REGION Network 13: ENCENDIDO ACTUADORES TUNEL 1
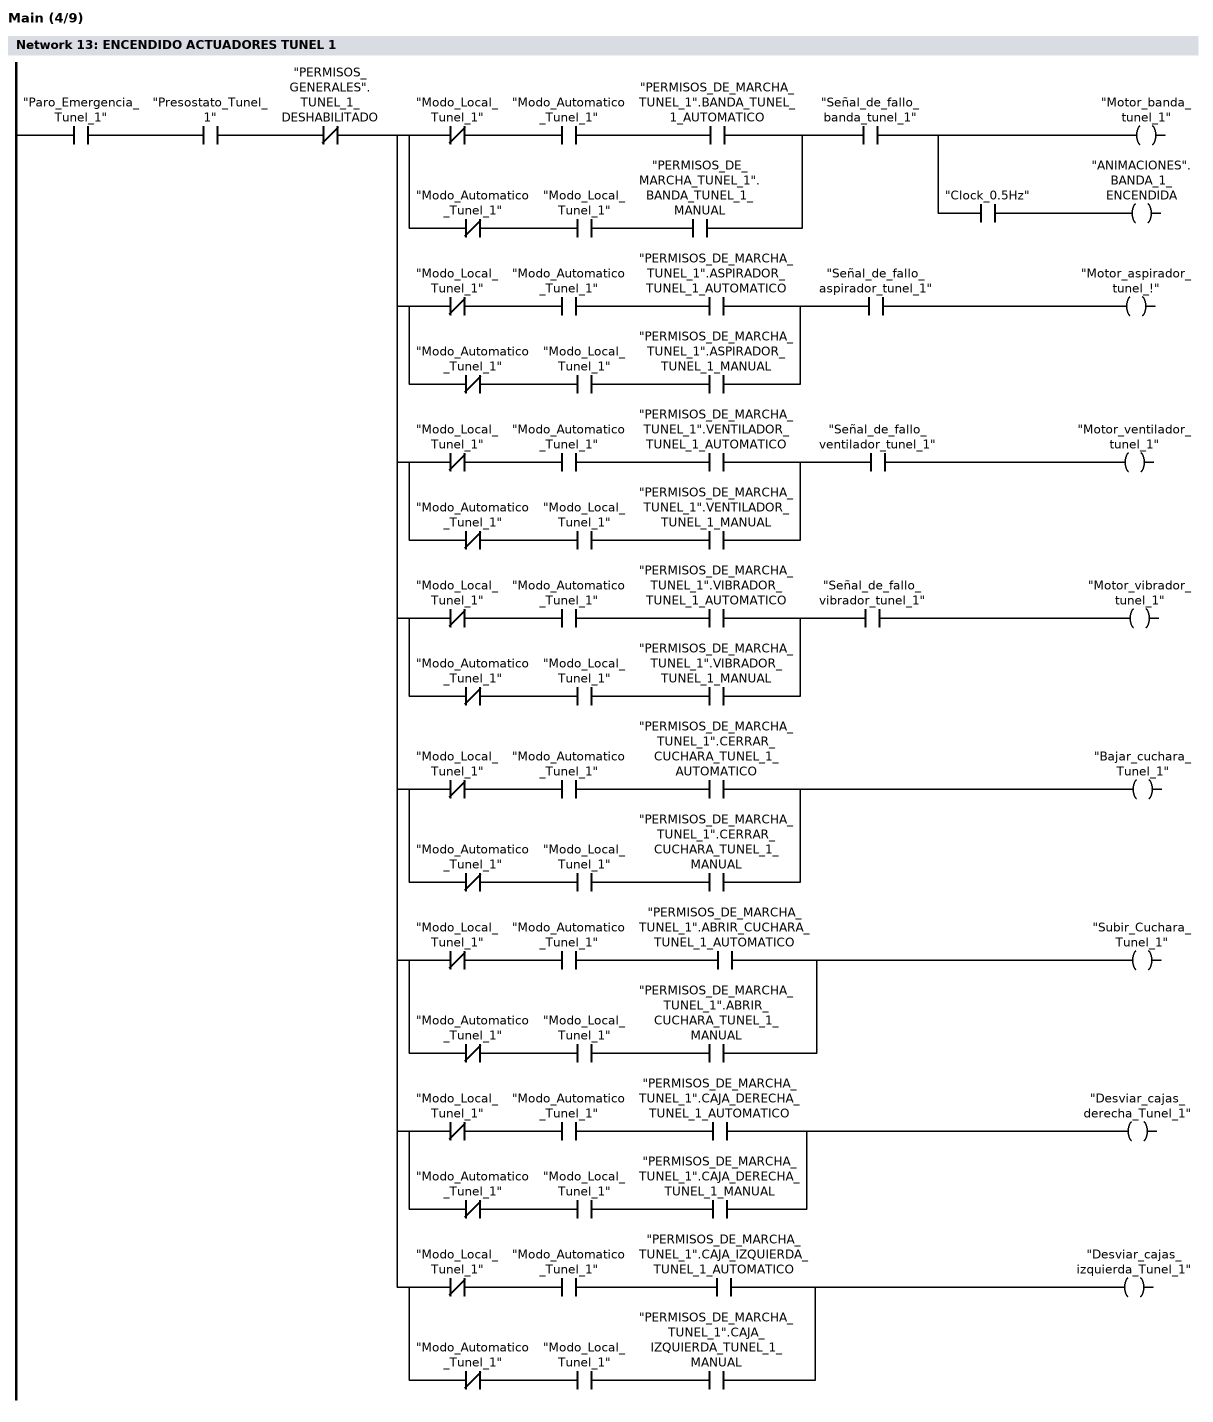
   RUNG wire#powerrail
      Contact( "Paro_Emergencia_Tunel_1" )
      Contact( "Presostato_Tunel_1" )
      I_Contact( "PERMISOS_GENERALES".TUNEL_1_DESHABILITADO )
      wire#w1
      I_Contact( "Modo_Local_Tunel_1" )
      Contact( "Modo_Automatico_Tunel_1" )
      Contact( "PERMISOS_DE_MARCHA_TUNEL_1".BANDA_TUNEL_1_AUTOMATICO )
      wire#w2
      Contact( "Señal_de_fallo_banda_tunel_1" )
      wire#w3
      Coil( "Motor_banda_tunel_1" )
   END_RUNG
   RUNG wire#w1
      I_Contact( "Modo_Automatico_Tunel_1" )
      Contact( "Modo_Local_Tunel_1" )
      Contact( "PERMISOS_DE_MARCHA_TUNEL_1".BANDA_TUNEL_1_MANUAL )
   END_RUNG wire#w2
   RUNG wire#w3
      Contact( "Clock_0.5Hz" )
      Coil( "ANIMACIONES".BANDA_1_ENCENDIDA )
   END_RUNG
   RUNG wire#w1
      I_Contact( "Modo_Local_Tunel_1" )
      Contact( "Modo_Automatico_Tunel_1" )
      Contact( "PERMISOS_DE_MARCHA_TUNEL_1".ASPIRADOR_TUNEL_1_AUTOMATICO )
      wire#w4
      Contact( "Señal_de_fallo_aspirador_tunel_1" )
      Coil( "Motor_aspirador_tunel_!" )
   END_RUNG
   RUNG wire#w1
      I_Contact( "Modo_Automatico_Tunel_1" )
      Contact( "Modo_Local_Tunel_1" )
      Contact( "PERMISOS_DE_MARCHA_TUNEL_1".ASPIRADOR_TUNEL_1_MANUAL )
   END_RUNG wire#w4
   RUNG wire#w1
      I_Contact( "Modo_Local_Tunel_1" )
      Contact( "Modo_Automatico_Tunel_1" )
      Contact( "PERMISOS_DE_MARCHA_TUNEL_1".VENTILADOR_TUNEL_1_AUTOMATICO )
      wire#w5
      Contact( "Señal_de_fallo_ventilador_tunel_1" )
      Coil( "Motor_ventilador_tunel_1" )
   END_RUNG
   RUNG wire#w1
      I_Contact( "Modo_Automatico_Tunel_1" )
      Contact( "Modo_Local_Tunel_1" )
      Contact( "PERMISOS_DE_MARCHA_TUNEL_1".VENTILADOR_TUNEL_1_MANUAL )
   END_RUNG wire#w5
   RUNG wire#w1
      I_Contact( "Modo_Local_Tunel_1" )
      Contact( "Modo_Automatico_Tunel_1" )
      Contact( "PERMISOS_DE_MARCHA_TUNEL_1".VIBRADOR_TUNEL_1_AUTOMATICO )
      wire#w6
      Contact( "Señal_de_fallo_vibrador_tunel_1" )
      Coil( "Motor_vibrador_tunel_1" )
   END_RUNG
   RUNG wire#w1
      I_Contact( "Modo_Automatico_Tunel_1" )
      Contact( "Modo_Local_Tunel_1" )
      Contact( "PERMISOS_DE_MARCHA_TUNEL_1".VIBRADOR_TUNEL_1_MANUAL )
   END_RUNG wire#w6
   RUNG wire#w1
      I_Contact( "Modo_Local_Tunel_1" )
      Contact( "Modo_Automatico_Tunel_1" )
      Contact( "PERMISOS_DE_MARCHA_TUNEL_1".CERRAR_CUCHARA_TUNEL_1_AUTOMATICO )
      wire#w7
      Coil( "Bajar_cuchara_Tunel_1" )
   END_RUNG
   RUNG wire#w1
      I_Contact( "Modo_Automatico_Tunel_1" )
      Contact( "Modo_Local_Tunel_1" )
      Contact( "PERMISOS_DE_MARCHA_TUNEL_1".CERRAR_CUCHARA_TUNEL_1_MANUAL )
   END_RUNG wire#w7
   RUNG wire#w1
      I_Contact( "Modo_Local_Tunel_1" )
      Contact( "Modo_Automatico_Tunel_1" )
      Contact( "PERMISOS_DE_MARCHA_TUNEL_1".ABRIR_CUCHARA_TUNEL_1_AUTOMATICO )
      wire#w8
      Coil( "Subir_Cuchara_Tunel_1" )
   END_RUNG
   RUNG wire#w1
      I_Contact( "Modo_Automatico_Tunel_1" )
      Contact( "Modo_Local_Tunel_1" )
      Contact( "PERMISOS_DE_MARCHA_TUNEL_1".ABRIR_CUCHARA_TUNEL_1_MANUAL )
   END_RUNG wire#w8
   RUNG wire#w1
      I_Contact( "Modo_Local_Tunel_1" )
      Contact( "Modo_Automatico_Tunel_1" )
      Contact( "PERMISOS_DE_MARCHA_TUNEL_1".CAJA_DERECHA_TUNEL_1_AUTOMATICO )
      wire#w9
      Coil( "Desviar_cajas_derecha_Tunel_1" )
   END_RUNG
   RUNG wire#w1
      I_Contact( "Modo_Automatico_Tunel_1" )
      Contact( "Modo_Local_Tunel_1" )
      Contact( "PERMISOS_DE_MARCHA_TUNEL_1".CAJA_DERECHA_TUNEL_1_MANUAL )
   END_RUNG wire#w9
   RUNG wire#w1
      I_Contact( "Modo_Local_Tunel_1" )
      Contact( "Modo_Automatico_Tunel_1" )
      Contact( "PERMISOS_DE_MARCHA_TUNEL_1".CAJA_IZQUIERDA_TUNEL_1_AUTOMATICO )
      wire#w10
      Coil( "Desviar_cajas_izquierda_Tunel_1" )
   END_RUNG
   RUNG wire#w1
      I_Contact( "Modo_Automatico_Tunel_1" )
      Contact( "Modo_Local_Tunel_1" )
      Contact( "PERMISOS_DE_MARCHA_TUNEL_1".CAJA_IZQUIERDA_TUNEL_1_MANUAL )
   END_RUNG wire#w10
   // the same network as SCL:
   #_w1 := "Paro_Emergencia_Tunel_1" AND "Presostato_Tunel_1" AND NOT "PERMISOS_GENERALES".TUNEL_1_DESHABILITADO;
   "Motor_banda_tunel_1" := #_w1 AND ((NOT "Modo_Local_Tunel_1" AND "Modo_Automatico_Tunel_1" AND "PERMISOS_DE_MARCHA_TUNEL_1".BANDA_TUNEL_1_AUTOMATICO) OR (NOT "Modo_Automatico_Tunel_1" AND "Modo_Local_Tunel_1" AND "PERMISOS_DE_MARCHA_TUNEL_1".BANDA_TUNEL_1_MANUAL)) AND "Señal_de_fallo_banda_tunel_1";
   "ANIMACIONES".BANDA_1_ENCENDIDA := "Motor_banda_tunel_1" AND "Clock_0.5Hz";
   "Motor_aspirador_tunel_!" := #_w1 AND ((NOT "Modo_Local_Tunel_1" AND "Modo_Automatico_Tunel_1" AND "PERMISOS_DE_MARCHA_TUNEL_1".ASPIRADOR_TUNEL_1_AUTOMATICO) OR (NOT "Modo_Automatico_Tunel_1" AND "Modo_Local_Tunel_1" AND "PERMISOS_DE_MARCHA_TUNEL_1".ASPIRADOR_TUNEL_1_MANUAL)) AND "Señal_de_fallo_aspirador_tunel_1";
   "Motor_ventilador_tunel_1" := #_w1 AND ((NOT "Modo_Local_Tunel_1" AND "Modo_Automatico_Tunel_1" AND "PERMISOS_DE_MARCHA_TUNEL_1".VENTILADOR_TUNEL_1_AUTOMATICO) OR (NOT "Modo_Automatico_Tunel_1" AND "Modo_Local_Tunel_1" AND "PERMISOS_DE_MARCHA_TUNEL_1".VENTILADOR_TUNEL_1_MANUAL)) AND "Señal_de_fallo_ventilador_tunel_1";
   "Motor_vibrador_tunel_1" := #_w1 AND ((NOT "Modo_Local_Tunel_1" AND "Modo_Automatico_Tunel_1" AND "PERMISOS_DE_MARCHA_TUNEL_1".VIBRADOR_TUNEL_1_AUTOMATICO) OR (NOT "Modo_Automatico_Tunel_1" AND "Modo_Local_Tunel_1" AND "PERMISOS_DE_MARCHA_TUNEL_1".VIBRADOR_TUNEL_1_MANUAL)) AND "Señal_de_fallo_vibrador_tunel_1";
   "Bajar_cuchara_Tunel_1" := #_w1 AND ((NOT "Modo_Local_Tunel_1" AND "Modo_Automatico_Tunel_1" AND "PERMISOS_DE_MARCHA_TUNEL_1".CERRAR_CUCHARA_TUNEL_1_AUTOMATICO) OR (NOT "Modo_Automatico_Tunel_1" AND "Modo_Local_Tunel_1" AND "PERMISOS_DE_MARCHA_TUNEL_1".CERRAR_CUCHARA_TUNEL_1_MANUAL));
   "Subir_Cuchara_Tunel_1" := #_w1 AND ((NOT "Modo_Local_Tunel_1" AND "Modo_Automatico_Tunel_1" AND "PERMISOS_DE_MARCHA_TUNEL_1".ABRIR_CUCHARA_TUNEL_1_AUTOMATICO) OR (NOT "Modo_Automatico_Tunel_1" AND "Modo_Local_Tunel_1" AND "PERMISOS_DE_MARCHA_TUNEL_1".ABRIR_CUCHARA_TUNEL_1_MANUAL));
   "Desviar_cajas_derecha_Tunel_1" := #_w1 AND ((NOT "Modo_Local_Tunel_1" AND "Modo_Automatico_Tunel_1" AND "PERMISOS_DE_MARCHA_TUNEL_1".CAJA_DERECHA_TUNEL_1_AUTOMATICO) OR (NOT "Modo_Automatico_Tunel_1" AND "Modo_Local_Tunel_1" AND "PERMISOS_DE_MARCHA_TUNEL_1".CAJA_DERECHA_TUNEL_1_MANUAL));
   "Desviar_cajas_izquierda_Tunel_1" := #_w1 AND ((NOT "Modo_Local_Tunel_1" AND "Modo_Automatico_Tunel_1" AND "PERMISOS_DE_MARCHA_TUNEL_1".CAJA_IZQUIERDA_TUNEL_1_AUTOMATICO) OR (NOT "Modo_Automatico_Tunel_1" AND "Modo_Local_Tunel_1" AND "PERMISOS_DE_MARCHA_TUNEL_1".CAJA_IZQUIERDA_TUNEL_1_MANUAL));
END_REGION

REGION Network 14: ENCENDIDO ACTUADORES TUNEL 2
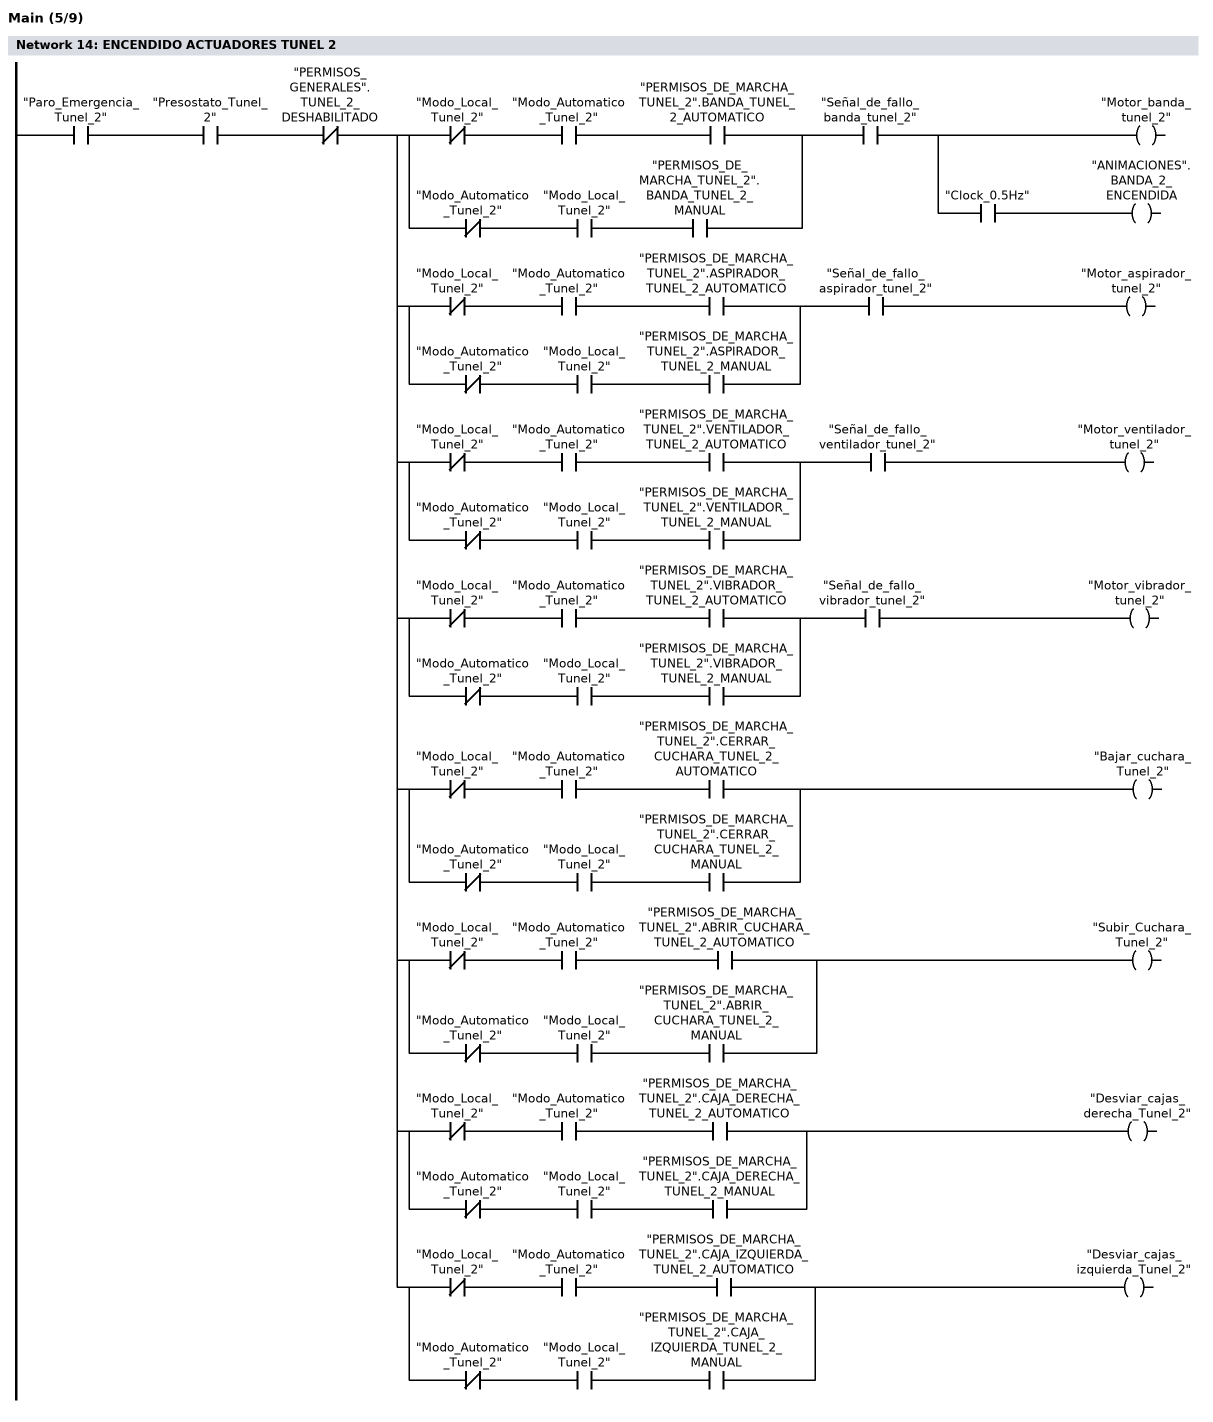
   RUNG wire#powerrail
      Contact( "Paro_Emergencia_Tunel_2" )
      Contact( "Presostato_Tunel_2" )
      I_Contact( "PERMISOS_GENERALES".TUNEL_2_DESHABILITADO )
      wire#w1
      I_Contact( "Modo_Local_Tunel_2" )
      Contact( "Modo_Automatico_Tunel_2" )
      Contact( "PERMISOS_DE_MARCHA_TUNEL_2".BANDA_TUNEL_2_AUTOMATICO )
      wire#w2
      Contact( "Señal_de_fallo_banda_tunel_2" )
      wire#w3
      Coil( "Motor_banda_tunel_2" )
   END_RUNG
   RUNG wire#w1
      I_Contact( "Modo_Automatico_Tunel_2" )
      Contact( "Modo_Local_Tunel_2" )
      Contact( "PERMISOS_DE_MARCHA_TUNEL_2".BANDA_TUNEL_2_MANUAL )
   END_RUNG wire#w2
   RUNG wire#w3
      Contact( "Clock_0.5Hz" )
      Coil( "ANIMACIONES".BANDA_2_ENCENDIDA )
   END_RUNG
   RUNG wire#w1
      I_Contact( "Modo_Local_Tunel_2" )
      Contact( "Modo_Automatico_Tunel_2" )
      Contact( "PERMISOS_DE_MARCHA_TUNEL_2".ASPIRADOR_TUNEL_2_AUTOMATICO )
      wire#w4
      Contact( "Señal_de_fallo_aspirador_tunel_2" )
      Coil( "Motor_aspirador_tunel_2" )
   END_RUNG
   RUNG wire#w1
      I_Contact( "Modo_Automatico_Tunel_2" )
      Contact( "Modo_Local_Tunel_2" )
      Contact( "PERMISOS_DE_MARCHA_TUNEL_2".ASPIRADOR_TUNEL_2_MANUAL )
   END_RUNG wire#w4
   RUNG wire#w1
      I_Contact( "Modo_Local_Tunel_2" )
      Contact( "Modo_Automatico_Tunel_2" )
      Contact( "PERMISOS_DE_MARCHA_TUNEL_2".VENTILADOR_TUNEL_2_AUTOMATICO )
      wire#w5
      Contact( "Señal_de_fallo_ventilador_tunel_2" )
      Coil( "Motor_ventilador_tunel_2" )
   END_RUNG
   RUNG wire#w1
      I_Contact( "Modo_Automatico_Tunel_2" )
      Contact( "Modo_Local_Tunel_2" )
      Contact( "PERMISOS_DE_MARCHA_TUNEL_2".VENTILADOR_TUNEL_2_MANUAL )
   END_RUNG wire#w5
   RUNG wire#w1
      I_Contact( "Modo_Local_Tunel_2" )
      Contact( "Modo_Automatico_Tunel_2" )
      Contact( "PERMISOS_DE_MARCHA_TUNEL_2".VIBRADOR_TUNEL_2_AUTOMATICO )
      wire#w6
      Contact( "Señal_de_fallo_vibrador_tunel_2" )
      Coil( "Motor_vibrador_tunel_2" )
   END_RUNG
   RUNG wire#w1
      I_Contact( "Modo_Automatico_Tunel_2" )
      Contact( "Modo_Local_Tunel_2" )
      Contact( "PERMISOS_DE_MARCHA_TUNEL_2".VIBRADOR_TUNEL_2_MANUAL )
   END_RUNG wire#w6
   RUNG wire#w1
      I_Contact( "Modo_Local_Tunel_2" )
      Contact( "Modo_Automatico_Tunel_2" )
      Contact( "PERMISOS_DE_MARCHA_TUNEL_2".CERRAR_CUCHARA_TUNEL_2_AUTOMATICO )
      wire#w7
      Coil( "Bajar_cuchara_Tunel_2" )
   END_RUNG
   RUNG wire#w1
      I_Contact( "Modo_Automatico_Tunel_2" )
      Contact( "Modo_Local_Tunel_2" )
      Contact( "PERMISOS_DE_MARCHA_TUNEL_2".CERRAR_CUCHARA_TUNEL_2_MANUAL )
   END_RUNG wire#w7
   RUNG wire#w1
      I_Contact( "Modo_Local_Tunel_2" )
      Contact( "Modo_Automatico_Tunel_2" )
      Contact( "PERMISOS_DE_MARCHA_TUNEL_2".ABRIR_CUCHARA_TUNEL_2_AUTOMATICO )
      wire#w8
      Coil( "Subir_Cuchara_Tunel_2" )
   END_RUNG
   RUNG wire#w1
      I_Contact( "Modo_Automatico_Tunel_2" )
      Contact( "Modo_Local_Tunel_2" )
      Contact( "PERMISOS_DE_MARCHA_TUNEL_2".ABRIR_CUCHARA_TUNEL_2_MANUAL )
   END_RUNG wire#w8
   RUNG wire#w1
      I_Contact( "Modo_Local_Tunel_2" )
      Contact( "Modo_Automatico_Tunel_2" )
      Contact( "PERMISOS_DE_MARCHA_TUNEL_2".CAJA_DERECHA_TUNEL_2_AUTOMATICO )
      wire#w9
      Coil( "Desviar_cajas_derecha_Tunel_2" )
   END_RUNG
   RUNG wire#w1
      I_Contact( "Modo_Automatico_Tunel_2" )
      Contact( "Modo_Local_Tunel_2" )
      Contact( "PERMISOS_DE_MARCHA_TUNEL_2".CAJA_DERECHA_TUNEL_2_MANUAL )
   END_RUNG wire#w9
   RUNG wire#w1
      I_Contact( "Modo_Local_Tunel_2" )
      Contact( "Modo_Automatico_Tunel_2" )
      Contact( "PERMISOS_DE_MARCHA_TUNEL_2".CAJA_IZQUIERDA_TUNEL_2_AUTOMATICO )
      wire#w10
      Coil( "Desviar_cajas_izquierda_Tunel_2" )
   END_RUNG
   RUNG wire#w1
      I_Contact( "Modo_Automatico_Tunel_2" )
      Contact( "Modo_Local_Tunel_2" )
      Contact( "PERMISOS_DE_MARCHA_TUNEL_2".CAJA_IZQUIERDA_TUNEL_2_MANUAL )
   END_RUNG wire#w10
   // the same network as SCL:
   #_w1 := "Paro_Emergencia_Tunel_2" AND "Presostato_Tunel_2" AND NOT "PERMISOS_GENERALES".TUNEL_2_DESHABILITADO;
   "Motor_banda_tunel_2" := #_w1 AND ((NOT "Modo_Local_Tunel_2" AND "Modo_Automatico_Tunel_2" AND "PERMISOS_DE_MARCHA_TUNEL_2".BANDA_TUNEL_2_AUTOMATICO) OR (NOT "Modo_Automatico_Tunel_2" AND "Modo_Local_Tunel_2" AND "PERMISOS_DE_MARCHA_TUNEL_2".BANDA_TUNEL_2_MANUAL)) AND "Señal_de_fallo_banda_tunel_2";
   "ANIMACIONES".BANDA_2_ENCENDIDA := "Motor_banda_tunel_2" AND "Clock_0.5Hz";
   "Motor_aspirador_tunel_2" := #_w1 AND ((NOT "Modo_Local_Tunel_2" AND "Modo_Automatico_Tunel_2" AND "PERMISOS_DE_MARCHA_TUNEL_2".ASPIRADOR_TUNEL_2_AUTOMATICO) OR (NOT "Modo_Automatico_Tunel_2" AND "Modo_Local_Tunel_2" AND "PERMISOS_DE_MARCHA_TUNEL_2".ASPIRADOR_TUNEL_2_MANUAL)) AND "Señal_de_fallo_aspirador_tunel_2";
   "Motor_ventilador_tunel_2" := #_w1 AND ((NOT "Modo_Local_Tunel_2" AND "Modo_Automatico_Tunel_2" AND "PERMISOS_DE_MARCHA_TUNEL_2".VENTILADOR_TUNEL_2_AUTOMATICO) OR (NOT "Modo_Automatico_Tunel_2" AND "Modo_Local_Tunel_2" AND "PERMISOS_DE_MARCHA_TUNEL_2".VENTILADOR_TUNEL_2_MANUAL)) AND "Señal_de_fallo_ventilador_tunel_2";
   "Motor_vibrador_tunel_2" := #_w1 AND ((NOT "Modo_Local_Tunel_2" AND "Modo_Automatico_Tunel_2" AND "PERMISOS_DE_MARCHA_TUNEL_2".VIBRADOR_TUNEL_2_AUTOMATICO) OR (NOT "Modo_Automatico_Tunel_2" AND "Modo_Local_Tunel_2" AND "PERMISOS_DE_MARCHA_TUNEL_2".VIBRADOR_TUNEL_2_MANUAL)) AND "Señal_de_fallo_vibrador_tunel_2";
   "Bajar_cuchara_Tunel_2" := #_w1 AND ((NOT "Modo_Local_Tunel_2" AND "Modo_Automatico_Tunel_2" AND "PERMISOS_DE_MARCHA_TUNEL_2".CERRAR_CUCHARA_TUNEL_2_AUTOMATICO) OR (NOT "Modo_Automatico_Tunel_2" AND "Modo_Local_Tunel_2" AND "PERMISOS_DE_MARCHA_TUNEL_2".CERRAR_CUCHARA_TUNEL_2_MANUAL));
   "Subir_Cuchara_Tunel_2" := #_w1 AND ((NOT "Modo_Local_Tunel_2" AND "Modo_Automatico_Tunel_2" AND "PERMISOS_DE_MARCHA_TUNEL_2".ABRIR_CUCHARA_TUNEL_2_AUTOMATICO) OR (NOT "Modo_Automatico_Tunel_2" AND "Modo_Local_Tunel_2" AND "PERMISOS_DE_MARCHA_TUNEL_2".ABRIR_CUCHARA_TUNEL_2_MANUAL));
   "Desviar_cajas_derecha_Tunel_2" := #_w1 AND ((NOT "Modo_Local_Tunel_2" AND "Modo_Automatico_Tunel_2" AND "PERMISOS_DE_MARCHA_TUNEL_2".CAJA_DERECHA_TUNEL_2_AUTOMATICO) OR (NOT "Modo_Automatico_Tunel_2" AND "Modo_Local_Tunel_2" AND "PERMISOS_DE_MARCHA_TUNEL_2".CAJA_DERECHA_TUNEL_2_MANUAL));
   "Desviar_cajas_izquierda_Tunel_2" := #_w1 AND ((NOT "Modo_Local_Tunel_2" AND "Modo_Automatico_Tunel_2" AND "PERMISOS_DE_MARCHA_TUNEL_2".CAJA_IZQUIERDA_TUNEL_2_AUTOMATICO) OR (NOT "Modo_Automatico_Tunel_2" AND "Modo_Local_Tunel_2" AND "PERMISOS_DE_MARCHA_TUNEL_2".CAJA_IZQUIERDA_TUNEL_2_MANUAL));
END_REGION

REGION Network 15: ENCENDIDO ACTUADORES TRANSPORTE
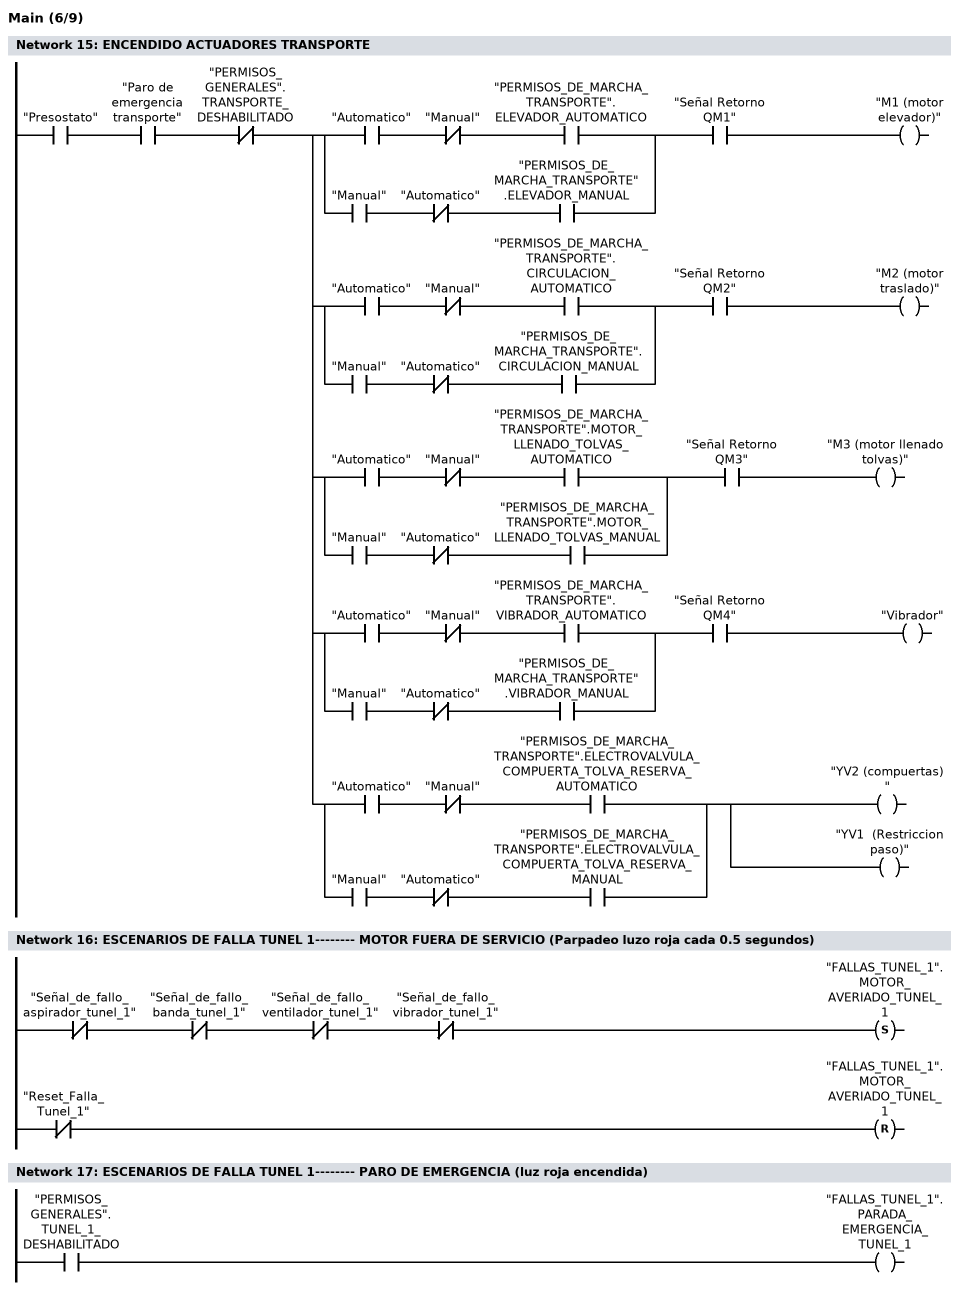
   RUNG wire#powerrail
      Contact( "Presostato" )
      Contact( "Paro de emergencia transporte" )
      I_Contact( "PERMISOS_GENERALES".TRANSPORTE_DESHABILITADO )
      wire#w1
      Contact( "Automatico" )
      I_Contact( "Manual" )
      Contact( "PERMISOS_DE_MARCHA_TRANSPORTE".ELEVADOR_AUTOMATICO )
      wire#w2
      Contact( "Señal Retorno QM1" )
      Coil( "M1 (motor elevador)" )
   END_RUNG
   RUNG wire#w1
      Contact( "Manual" )
      I_Contact( "Automatico" )
      Contact( "PERMISOS_DE_MARCHA_TRANSPORTE".ELEVADOR_MANUAL )
   END_RUNG wire#w2
   RUNG wire#w1
      Contact( "Automatico" )
      I_Contact( "Manual" )
      Contact( "PERMISOS_DE_MARCHA_TRANSPORTE".CIRCULACION_AUTOMATICO )
      wire#w3
      Contact( "Señal Retorno QM2" )
      Coil( "M2 (motor traslado)" )
   END_RUNG
   RUNG wire#w1
      Contact( "Manual" )
      I_Contact( "Automatico" )
      Contact( "PERMISOS_DE_MARCHA_TRANSPORTE".CIRCULACION_MANUAL )
   END_RUNG wire#w3
   RUNG wire#w1
      Contact( "Automatico" )
      I_Contact( "Manual" )
      Contact( "PERMISOS_DE_MARCHA_TRANSPORTE".MOTOR_LLENADO_TOLVAS_AUTOMATICO )
      wire#w4
      Contact( "Señal Retorno QM3" )
      Coil( "M3 (motor llenado tolvas)" )
   END_RUNG
   RUNG wire#w1
      Contact( "Manual" )
      I_Contact( "Automatico" )
      Contact( "PERMISOS_DE_MARCHA_TRANSPORTE".MOTOR_LLENADO_TOLVAS_MANUAL )
   END_RUNG wire#w4
   RUNG wire#w1
      Contact( "Automatico" )
      I_Contact( "Manual" )
      Contact( "PERMISOS_DE_MARCHA_TRANSPORTE".VIBRADOR_AUTOMATICO )
      wire#w5
      Contact( "Señal Retorno QM4" )
      Coil( "Vibrador" )
   END_RUNG
   RUNG wire#w1
      Contact( "Manual" )
      I_Contact( "Automatico" )
      Contact( "PERMISOS_DE_MARCHA_TRANSPORTE".VIBRADOR_MANUAL )
   END_RUNG wire#w5
   RUNG wire#w1
      Contact( "Automatico" )
      I_Contact( "Manual" )
      Contact( "PERMISOS_DE_MARCHA_TRANSPORTE".ELECTROVALVULA_COMPUERTA_TOLVA_RESERVA_AUTOMATICO )
      wire#w6
      Coil( "YV2 (compuertas)" )
   END_RUNG
   RUNG wire#w1
      Contact( "Manual" )
      I_Contact( "Automatico" )
      Contact( "PERMISOS_DE_MARCHA_TRANSPORTE".ELECTROVALVULA_COMPUERTA_TOLVA_RESERVA_MANUAL )
   END_RUNG wire#w6
   RUNG wire#w6
      Coil( "YV1  (Restriccion paso)" )
   END_RUNG
   // the same network as SCL:
   #_w1 := "Presostato" AND "Paro de emergencia transporte" AND NOT "PERMISOS_GENERALES".TRANSPORTE_DESHABILITADO;
   "M1 (motor elevador)" := #_w1 AND (("Automatico" AND NOT "Manual" AND "PERMISOS_DE_MARCHA_TRANSPORTE".ELEVADOR_AUTOMATICO) OR ("Manual" AND NOT "Automatico" AND "PERMISOS_DE_MARCHA_TRANSPORTE".ELEVADOR_MANUAL)) AND "Señal Retorno QM1";
   "M2 (motor traslado)" := #_w1 AND (("Automatico" AND NOT "Manual" AND "PERMISOS_DE_MARCHA_TRANSPORTE".CIRCULACION_AUTOMATICO) OR ("Manual" AND NOT "Automatico" AND "PERMISOS_DE_MARCHA_TRANSPORTE".CIRCULACION_MANUAL)) AND "Señal Retorno QM2";
   "M3 (motor llenado tolvas)" := #_w1 AND (("Automatico" AND NOT "Manual" AND "PERMISOS_DE_MARCHA_TRANSPORTE".MOTOR_LLENADO_TOLVAS_AUTOMATICO) OR ("Manual" AND NOT "Automatico" AND "PERMISOS_DE_MARCHA_TRANSPORTE".MOTOR_LLENADO_TOLVAS_MANUAL)) AND "Señal Retorno QM3";
   "Vibrador" := #_w1 AND (("Automatico" AND NOT "Manual" AND "PERMISOS_DE_MARCHA_TRANSPORTE".VIBRADOR_AUTOMATICO) OR ("Manual" AND NOT "Automatico" AND "PERMISOS_DE_MARCHA_TRANSPORTE".VIBRADOR_MANUAL)) AND "Señal Retorno QM4";
   "YV2 (compuertas)" := #_w1 AND (("Automatico" AND NOT "Manual" AND "PERMISOS_DE_MARCHA_TRANSPORTE".ELECTROVALVULA_COMPUERTA_TOLVA_RESERVA_AUTOMATICO) OR ("Manual" AND NOT "Automatico" AND "PERMISOS_DE_MARCHA_TRANSPORTE".ELECTROVALVULA_COMPUERTA_TOLVA_RESERVA_MANUAL));
   "YV1  (Restriccion paso)" := "YV2 (compuertas)";
END_REGION

REGION Network 16: ESCENARIOS DE FALLA TUNEL 1-------- MOTOR FUERA DE SERVICIO (Parpadeo luzo roja cada 0.5 segundos)
   RUNG wire#powerrail
      I_Contact( "Señal_de_fallo_aspirador_tunel_1" )
      I_Contact( "Señal_de_fallo_banda_tunel_1" )
      I_Contact( "Señal_de_fallo_ventilador_tunel_1" )
      I_Contact( "Señal_de_fallo_vibrador_tunel_1" )
      S_Coil( "FALLAS_TUNEL_1".MOTOR_AVERIADO_TUNEL_1 )
   END_RUNG
   RUNG wire#powerrail
      I_Contact( "Reset_Falla_Tunel_1" )
      R_Coil( "FALLAS_TUNEL_1".MOTOR_AVERIADO_TUNEL_1 )
   END_RUNG
   // the same network as SCL:
   IF NOT "Señal_de_fallo_aspirador_tunel_1" AND NOT "Señal_de_fallo_banda_tunel_1" AND NOT "Señal_de_fallo_ventilador_tunel_1" AND NOT "Señal_de_fallo_vibrador_tunel_1" THEN
       "FALLAS_TUNEL_1".MOTOR_AVERIADO_TUNEL_1 := TRUE;
   END_IF;
   IF NOT "Reset_Falla_Tunel_1" THEN "FALLAS_TUNEL_1".MOTOR_AVERIADO_TUNEL_1 := FALSE; END_IF;
END_REGION

REGION Network 17: ESCENARIOS DE FALLA TUNEL 1-------- PARO DE EMERGENCIA (luz roja encendida)
   RUNG wire#powerrail
      Contact( "PERMISOS_GENERALES".TUNEL_1_DESHABILITADO )
      Coil( "FALLAS_TUNEL_1".PARADA_EMERGENCIA_TUNEL_1 )
   END_RUNG
   // the same network as SCL:
   "FALLAS_TUNEL_1".PARADA_EMERGENCIA_TUNEL_1 := "PERMISOS_GENERALES".TUNEL_1_DESHABILITADO;
END_REGION

REGION Network 18: ENCENDIDO LAMPARA ROJA TUNEL 1
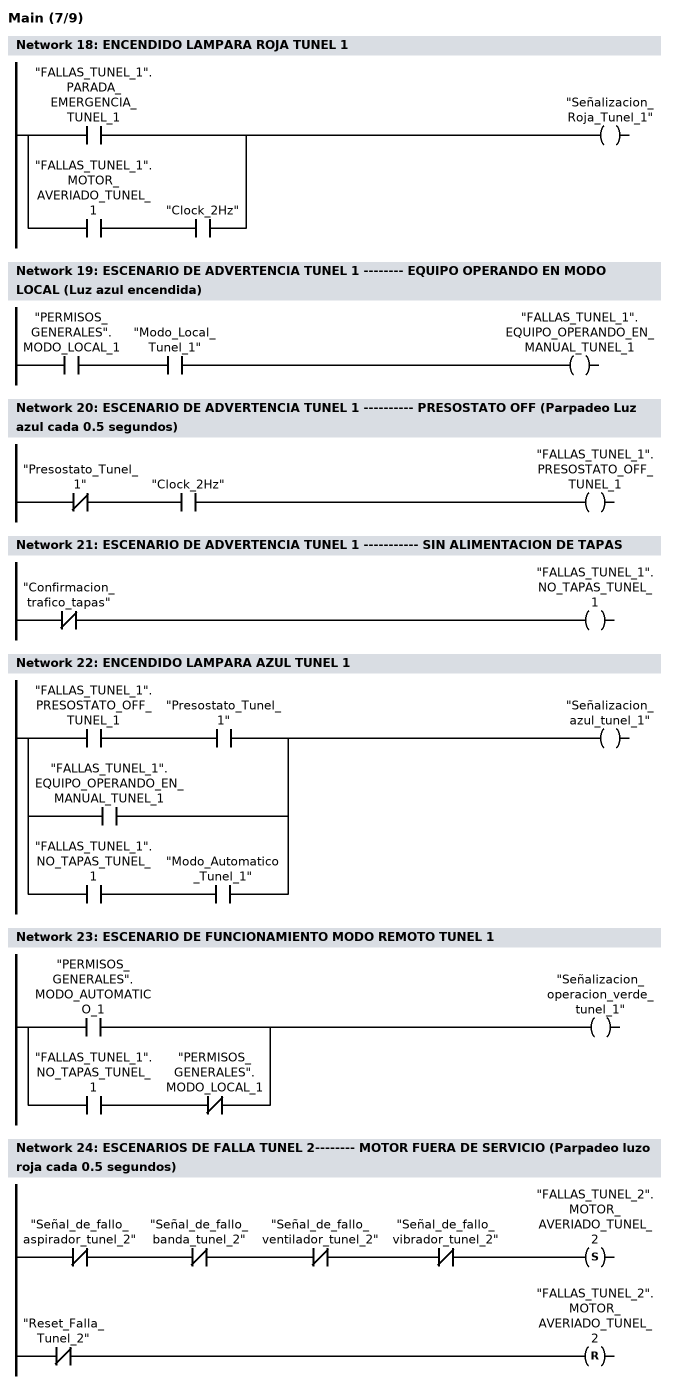
   RUNG wire#powerrail
      Contact( "FALLAS_TUNEL_1".PARADA_EMERGENCIA_TUNEL_1 )
      wire#w1
      Coil( "Señalizacion_Roja_Tunel_1" )
   END_RUNG
   RUNG wire#powerrail
      Contact( "FALLAS_TUNEL_1".MOTOR_AVERIADO_TUNEL_1 )
      Contact( "Clock_2Hz" )
   END_RUNG wire#w1
   // the same network as SCL:
   "Señalizacion_Roja_Tunel_1" := "FALLAS_TUNEL_1".PARADA_EMERGENCIA_TUNEL_1 OR ("FALLAS_TUNEL_1".MOTOR_AVERIADO_TUNEL_1 AND "Clock_2Hz");
END_REGION

REGION Network 19: ESCENARIO DE ADVERTENCIA TUNEL 1 -------- EQUIPO OPERANDO EN MODO LOCAL (Luz azul encendida)
   RUNG wire#powerrail
      Contact( "PERMISOS_GENERALES".MODO_LOCAL_1 )
      Contact( "Modo_Local_Tunel_1" )
      Coil( "FALLAS_TUNEL_1".EQUIPO_OPERANDO_EN_MANUAL_TUNEL_1 )
   END_RUNG
   // the same network as SCL:
   "FALLAS_TUNEL_1".EQUIPO_OPERANDO_EN_MANUAL_TUNEL_1 := "PERMISOS_GENERALES".MODO_LOCAL_1 AND "Modo_Local_Tunel_1";
END_REGION

REGION Network 20: ESCENARIO DE ADVERTENCIA TUNEL 1 ---------- PRESOSTATO OFF (Parpadeo Luz azul cada 0.5 segundos)
   RUNG wire#powerrail
      I_Contact( "Presostato_Tunel_1" )
      Contact( "Clock_2Hz" )
      Coil( "FALLAS_TUNEL_1".PRESOSTATO_OFF_TUNEL_1 )
   END_RUNG
   // the same network as SCL:
   "FALLAS_TUNEL_1".PRESOSTATO_OFF_TUNEL_1 := NOT "Presostato_Tunel_1" AND "Clock_2Hz";
END_REGION

REGION Network 21: ESCENARIO DE ADVERTENCIA TUNEL 1 ----------- SIN ALIMENTACION DE TAPAS
   RUNG wire#powerrail
      I_Contact( "Confirmacion_trafico_tapas" )
      Coil( "FALLAS_TUNEL_1".NO_TAPAS_TUNEL_1 )
   END_RUNG
   // the same network as SCL:
   "FALLAS_TUNEL_1".NO_TAPAS_TUNEL_1 := NOT "Confirmacion_trafico_tapas";
END_REGION

REGION Network 22: ENCENDIDO LAMPARA AZUL TUNEL 1
   RUNG wire#powerrail
      Contact( "FALLAS_TUNEL_1".PRESOSTATO_OFF_TUNEL_1 )
      Contact( "Presostato_Tunel_1" )
      wire#w1
      Coil( "Señalizacion_azul_tunel_1" )
   END_RUNG
   RUNG wire#powerrail
      Contact( "FALLAS_TUNEL_1".EQUIPO_OPERANDO_EN_MANUAL_TUNEL_1 )
   END_RUNG wire#w1
   RUNG wire#powerrail
      Contact( "FALLAS_TUNEL_1".NO_TAPAS_TUNEL_1 )
      Contact( "Modo_Automatico_Tunel_1" )
   END_RUNG wire#w1
   // the same network as SCL:
   "Señalizacion_azul_tunel_1" := ("FALLAS_TUNEL_1".PRESOSTATO_OFF_TUNEL_1 AND "Presostato_Tunel_1") OR "FALLAS_TUNEL_1".EQUIPO_OPERANDO_EN_MANUAL_TUNEL_1 OR ("FALLAS_TUNEL_1".NO_TAPAS_TUNEL_1 AND "Modo_Automatico_Tunel_1");
END_REGION

REGION Network 23: ESCENARIO DE FUNCIONAMIENTO MODO REMOTO TUNEL 1
   RUNG wire#powerrail
      Contact( "PERMISOS_GENERALES".MODO_AUTOMATICO_1 )
      wire#w1
      Coil( "Señalizacion_operacion_verde_tunel_1" )
   END_RUNG
   RUNG wire#powerrail
      Contact( "FALLAS_TUNEL_1".NO_TAPAS_TUNEL_1 )
      I_Contact( "PERMISOS_GENERALES".MODO_LOCAL_1 )
   END_RUNG wire#w1
   // the same network as SCL:
   "Señalizacion_operacion_verde_tunel_1" := "PERMISOS_GENERALES".MODO_AUTOMATICO_1 OR ("FALLAS_TUNEL_1".NO_TAPAS_TUNEL_1 AND NOT "PERMISOS_GENERALES".MODO_LOCAL_1);
END_REGION

REGION Network 24: ESCENARIOS DE FALLA TUNEL 2-------- MOTOR FUERA DE SERVICIO (Parpadeo luzo roja cada 0.5 segundos)
   RUNG wire#powerrail
      I_Contact( "Señal_de_fallo_aspirador_tunel_2" )
      I_Contact( "Señal_de_fallo_banda_tunel_2" )
      I_Contact( "Señal_de_fallo_ventilador_tunel_2" )
      I_Contact( "Señal_de_fallo_vibrador_tunel_2" )
      S_Coil( "FALLAS_TUNEL_2".MOTOR_AVERIADO_TUNEL_2 )
   END_RUNG
   RUNG wire#powerrail
      I_Contact( "Reset_Falla_Tunel_2" )
      R_Coil( "FALLAS_TUNEL_2".MOTOR_AVERIADO_TUNEL_2 )
   END_RUNG
   // the same network as SCL:
   IF NOT "Señal_de_fallo_aspirador_tunel_2" AND NOT "Señal_de_fallo_banda_tunel_2" AND NOT "Señal_de_fallo_ventilador_tunel_2" AND NOT "Señal_de_fallo_vibrador_tunel_2" THEN
       "FALLAS_TUNEL_2".MOTOR_AVERIADO_TUNEL_2 := TRUE;
   END_IF;
   IF NOT "Reset_Falla_Tunel_2" THEN "FALLAS_TUNEL_2".MOTOR_AVERIADO_TUNEL_2 := FALSE; END_IF;
END_REGION

REGION Network 25: ESCENARIOS DE FALLA TUNEL 2-------- PARO DE EMERGENCIA (luz roja encendida)
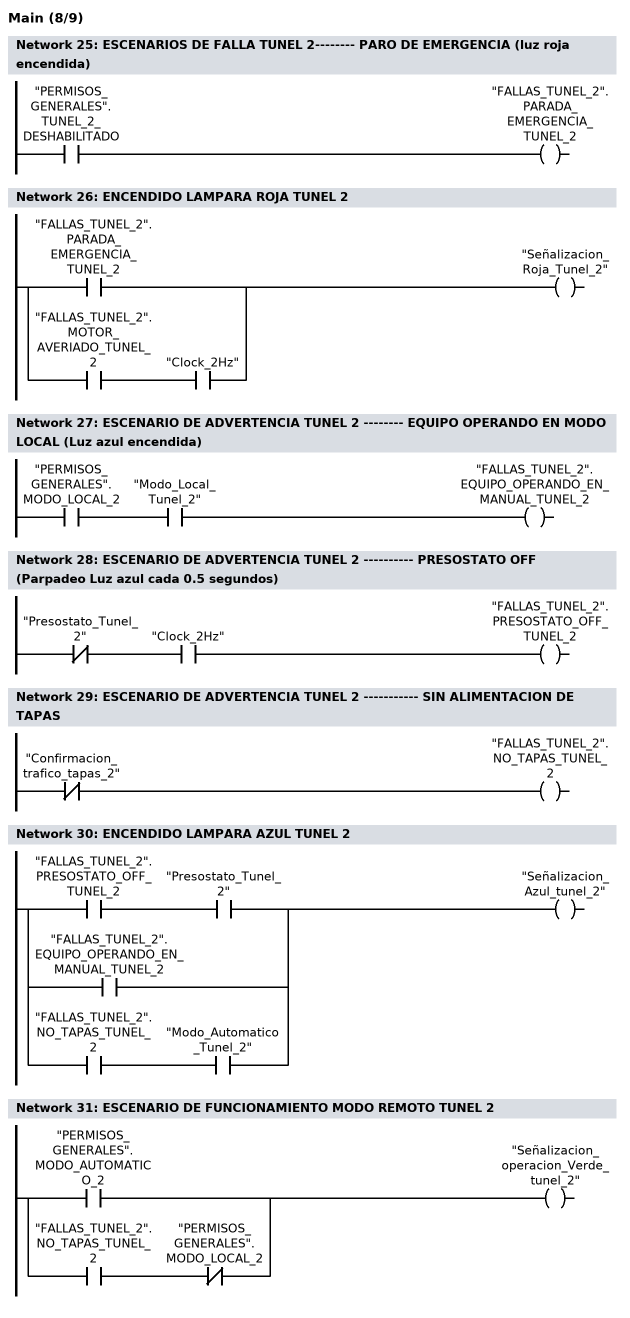
   RUNG wire#powerrail
      Contact( "PERMISOS_GENERALES".TUNEL_2_DESHABILITADO )
      Coil( "FALLAS_TUNEL_2".PARADA_EMERGENCIA_TUNEL_2 )
   END_RUNG
   // the same network as SCL:
   "FALLAS_TUNEL_2".PARADA_EMERGENCIA_TUNEL_2 := "PERMISOS_GENERALES".TUNEL_2_DESHABILITADO;
END_REGION

REGION Network 26: ENCENDIDO LAMPARA ROJA TUNEL 2
   RUNG wire#powerrail
      Contact( "FALLAS_TUNEL_2".PARADA_EMERGENCIA_TUNEL_2 )
      wire#w1
      Coil( "Señalizacion_Roja_Tunel_2" )
   END_RUNG
   RUNG wire#powerrail
      Contact( "FALLAS_TUNEL_2".MOTOR_AVERIADO_TUNEL_2 )
      Contact( "Clock_2Hz" )
   END_RUNG wire#w1
   // the same network as SCL:
   "Señalizacion_Roja_Tunel_2" := "FALLAS_TUNEL_2".PARADA_EMERGENCIA_TUNEL_2 OR ("FALLAS_TUNEL_2".MOTOR_AVERIADO_TUNEL_2 AND "Clock_2Hz");
END_REGION

REGION Network 27: ESCENARIO DE ADVERTENCIA TUNEL 2 -------- EQUIPO OPERANDO EN MODO LOCAL (Luz azul encendida)
   RUNG wire#powerrail
      Contact( "PERMISOS_GENERALES".MODO_LOCAL_2 )
      Contact( "Modo_Local_Tunel_2" )
      Coil( "FALLAS_TUNEL_2".EQUIPO_OPERANDO_EN_MANUAL_TUNEL_2 )
   END_RUNG
   // the same network as SCL:
   "FALLAS_TUNEL_2".EQUIPO_OPERANDO_EN_MANUAL_TUNEL_2 := "PERMISOS_GENERALES".MODO_LOCAL_2 AND "Modo_Local_Tunel_2";
END_REGION

REGION Network 28: ESCENARIO DE ADVERTENCIA TUNEL 2 ---------- PRESOSTATO OFF (Parpadeo Luz azul cada 0.5 segundos)
   RUNG wire#powerrail
      I_Contact( "Presostato_Tunel_2" )
      Contact( "Clock_2Hz" )
      Coil( "FALLAS_TUNEL_2".PRESOSTATO_OFF_TUNEL_2 )
   END_RUNG
   // the same network as SCL:
   "FALLAS_TUNEL_2".PRESOSTATO_OFF_TUNEL_2 := NOT "Presostato_Tunel_2" AND "Clock_2Hz";
END_REGION

REGION Network 29: ESCENARIO DE ADVERTENCIA TUNEL 2 ----------- SIN ALIMENTACION DE TAPAS
   RUNG wire#powerrail
      I_Contact( "Confirmacion_trafico_tapas_2" )
      Coil( "FALLAS_TUNEL_2".NO_TAPAS_TUNEL_2 )
   END_RUNG
   // the same network as SCL:
   "FALLAS_TUNEL_2".NO_TAPAS_TUNEL_2 := NOT "Confirmacion_trafico_tapas_2";
END_REGION

REGION Network 30: ENCENDIDO LAMPARA AZUL TUNEL 2
   RUNG wire#powerrail
      Contact( "FALLAS_TUNEL_2".PRESOSTATO_OFF_TUNEL_2 )
      Contact( "Presostato_Tunel_2" )
      wire#w1
      Coil( "Señalizacion_Azul_tunel_2" )
   END_RUNG
   RUNG wire#powerrail
      Contact( "FALLAS_TUNEL_2".EQUIPO_OPERANDO_EN_MANUAL_TUNEL_2 )
   END_RUNG wire#w1
   RUNG wire#powerrail
      Contact( "FALLAS_TUNEL_2".NO_TAPAS_TUNEL_2 )
      Contact( "Modo_Automatico_Tunel_2" )
   END_RUNG wire#w1
   // the same network as SCL:
   "Señalizacion_Azul_tunel_2" := ("FALLAS_TUNEL_2".PRESOSTATO_OFF_TUNEL_2 AND "Presostato_Tunel_2") OR "FALLAS_TUNEL_2".EQUIPO_OPERANDO_EN_MANUAL_TUNEL_2 OR ("FALLAS_TUNEL_2".NO_TAPAS_TUNEL_2 AND "Modo_Automatico_Tunel_2");
END_REGION

REGION Network 31: ESCENARIO DE FUNCIONAMIENTO MODO REMOTO TUNEL 2
   RUNG wire#powerrail
      Contact( "PERMISOS_GENERALES".MODO_AUTOMATICO_2 )
      wire#w1
      Coil( "Señalizacion_operacion_Verde_tunel_2" )
   END_RUNG
   RUNG wire#powerrail
      Contact( "FALLAS_TUNEL_2".NO_TAPAS_TUNEL_2 )
      I_Contact( "PERMISOS_GENERALES".MODO_LOCAL_2 )
   END_RUNG wire#w1
   // the same network as SCL:
   "Señalizacion_operacion_Verde_tunel_2" := "PERMISOS_GENERALES".MODO_AUTOMATICO_2 OR ("FALLAS_TUNEL_2".NO_TAPAS_TUNEL_2 AND NOT "PERMISOS_GENERALES".MODO_LOCAL_2);
END_REGION

REGION Network 32: ANIMACIONES TUNEL_1